   "Carrier_35_PB3_ProdHoldRH" AT %I2117.2 : Bool;   // PB 3 PRODUCTION HOLD RH
   "Carrier_35_PB4_ResetRH" AT %I2117.3 : Bool;   // PB 4 RESET RH
   "Carrier_35_SpareInput(4_14)" AT %I2117.4 : Bool;   // SPARE INPUT
   "Carrier_35_SpareInput(4_15)" AT %I2117.5 : Bool;   // SPARE INPUT
   "Carrier_35_SpareInput(4_16)" AT %I2117.6 : Bool;   // SPARE INPUT
   "Carrier_35_SpareInput(4_17)" AT %I2117.7 : Bool;   // SPARE INPUT
   "Carrier_35_Slot5_Output" AT %IW2118 : Word;   // SLOT 5 OUTPUT WORD
   "Carrier_35_IRD400_HMI_24VDC_ENABLE" AT %I2118.0 : Bool;   // IRD 400 PANEL HMI 24V DC POWER
   "Carrier_35_FaultLight_LH" AT %I2118.1 : Bool;   // FAULT LIGHT LH
   "Carrier_35_RunLight_LH" AT %I2118.2 : Bool;   // RUN LIGHT LH
   "Carrier_35_FaultLight_RH" AT %I2118.3 : Bool;   // FAULT LIGHT RH
   "Carrier_35_RunLight_RH" AT %I2118.4 : Bool;   // RUN LIGHT RH
   "Carrier_35_SpareOutput(5_5)" AT %I2118.5 : Bool;   // SPARE OUTPUT
   "Carrier_35_SpareOutput(5_6)" AT %I2118.6 : Bool;   // SPARE OUTPUT
   "Carrier_35_SpareOutput(5_7)" AT %I2118.7 : Bool;   // SPARE OUTPUT
   "Carrier_35_ActualSpeed" AT %IW2120 : Word;   // ACTUAL SPEED
   "Carrier_35_CarrierDriveAlarm" AT %IW2122 : Word;   // CARRIER DRIVE ALARM
   "Carrier_35_CarrierDriveWarning" AT %IW2124 : Word;   // CARRIER DRIVE WARNING
   "Carrier_36_Status" AT %IW2150 : Word;   // CARRIER STATUS WORD
   "Carrier_36_Status.0" AT %I2150.0 : Bool;   // HEARTBEAT
   "Carrier_36_Status.1" AT %I2150.1 : Bool;   // MANUAL
   "Carrier_36_Status.2" AT %I2150.2 : Bool;   // IN_AUTO
   "Carrier_36_Status.3" AT %I2150.3 : Bool;   // POSITIONING_COMPLETE
   "Carrier_36_Status.4" AT %I2150.4 : Bool;   // PRODUCTION HOLD
   "Carrier_36_Status.5" AT %I2150.5 : Bool;   // CARRIER MOVING FORWARD
   "Carrier_36_Status.6" AT %I2150.6 : Bool;   // CARRIER MOVING REVERSE
   "Carrier_36_Status.7" AT %I2150.7 : Bool;   // CARRIER FAULT
   "Carrier_36_Status.8" AT %I2151.0 : Bool;   // CRASH DETECT TRIPPED
   "Carrier_36_Status.9" AT %I2151.1 : Bool;
   "Carrier_36_Status.10" AT %I2151.2 : Bool;
   "Carrier_36_Status.11" AT %I2151.3 : Bool;
   "Carrier_36_Status.12" AT %I2151.4 : Bool;
   "Carrier_36_Status.13" AT %I2151.5 : Bool;
   "Carrier_36_Status.14" AT %I2151.6 : Bool;
   "Carrier_36_Status.15" AT %I2151.7 : Bool;
   "Carrier_36_SDCFaultCode" AT %IW2152 : Word;   // SDC FAULT CODE
   "Carrier_36_CarrierPosition" AT %ID2154 : DWord;   // CARRIER POSITION
   "Carrier_36_CarrierNumber" AT %IW2158 : Word;   // CARRIER NUMBER
   "Carrier_36_G120DControlWord" AT %IW2160 : Word;   // G120D_STW1_CONTROL
   "Carrier_36_G120DControlWord.0" AT %I2160.0 : Bool;   // Bit_00_ON
   "Carrier_36_G120DControlWord.1" AT %I2160.1 : Bool;   // Bit_01_AUS2_INH
   "Carrier_36_G120DControlWord.2" AT %I2160.2 : Bool;   // Bit_02_AUS3_STOP
   "Carrier_36_G120DControlWord.3" AT %I2160.3 : Bool;   // Bit_03_EN
   "Carrier_36_G120DControlWord.4" AT %I2160.4 : Bool;   // Bit_04_EN_RAMP
   "Carrier_36_G120DControlWord.5" AT %I2160.5 : Bool;   // Bit_05_START_RAMP
   "Carrier_36_G120DControlWord.6" AT %I2160.6 : Bool;   // Bit_06_SETPOINT
   "Carrier_36_G120DControlWord.7" AT %I2160.7 : Bool;   // Bit_07_RESET
   "Carrier_36_G120DControlWord.8" AT %I2161.0 : Bool;   // Bit_08_JOG_R
   "Carrier_36_G120DControlWord.9" AT %I2161.1 : Bool;   // Bit_09_JOG_L
   "Carrier_36_G120DControlWord.10" AT %I2161.2 : Bool;   // Bit_10_CONTR_PLC
   "Carrier_36_G120DControlWord.11" AT %I2161.3 : Bool;   // Bit_11_REVERSE
   "Carrier_36_G120DControlWord.12" AT %I2161.4 : Bool;   // Bit_12_BRAKE_RELEASE
   "Carrier_36_G120DControlWord.13" AT %I2161.5 : Bool;   // Bit_13_DDS
   "Carrier_36_G120DControlWord.14" AT %I2161.6 : Bool;   // Bit_14_DO0
   "Carrier_36_G120DControlWord.15" AT %I2161.7 : Bool;   // Bit_15_DO1
   "Carrier_36_G120DStatusWord" AT %IW2162 : Word;   // G120D_ZSW1_STATUS
   "Carrier_36_G120DStatusWord.0" AT %I2162.0 : Bool;   // Bit_00_READY_RUN
   "Carrier_36_G120DStatusWord.1" AT %I2162.1 : Bool;   // Bit_01_READY_ON
   "Carrier_36_G120DStatusWord.2" AT %I2162.2 : Bool;   // Bit_02_ENABLE
   "Carrier_36_G120DStatusWord.3" AT %I2162.3 : Bool;   // Bit_03_FAULT
   "Carrier_36_G120DStatusWord.4" AT %I2162.4 : Bool;   // Bit_04_OFF2
   "Carrier_36_G120DStatusWord.5" AT %I2162.5 : Bool;   // Bit_05_OFF3
   "Carrier_36_G120DStatusWord.6" AT %I2162.6 : Bool;   // Bit_06_LOCK_OUT
   "Carrier_36_G120DStatusWord.7" AT %I2162.7 : Bool;   // Bit_07_WARN
   "Carrier_36_G120DStatusWord.8" AT %I2163.0 : Bool;   // Bit_08_NO_DEVIATION
   "Carrier_36_G120DStatusWord.9" AT %I2163.1 : Bool;   // Bit_09_CONTR_PLC
   "Carrier_36_G120DStatusWord.10" AT %I2163.2 : Bool;   // Bit_10_F_MAX
   "Carrier_36_G120DStatusWord.11" AT %I2163.3 : Bool;   // Bit_11_LIMIT_REACHED
   "Carrier_36_G120DStatusWord.12" AT %I2163.4 : Bool;   // Bit_12_BRAKE_OPEN
   "Carrier_36_G120DStatusWord.13" AT %I2163.5 : Bool;   // Bit_13_NO_OVERTEMP
   "Carrier_36_G120DStatusWord.14" AT %I2163.6 : Bool;   // Bit_14_CW_CCW
   "Carrier_36_G120DStatusWord.15" AT %I2163.7 : Bool;   // Bit_15_OVERL
   "Carrier_36_Slot2_Input" AT %IW2164 : Word;   // SLOT 2 INPUT WORD
   "Carrier_36_CrashDetectSW" AT %I2164.0 : Bool;   // CRASH DETECT SW
   "Carrier_36_SpareSafetyInput(2_1)" AT %I2164.1 : Bool;   // SPARE SAFETY INPUT
   "Carrier_36_SpareSafetyInput(2_2)" AT %I2164.2 : Bool;   // SPARE SAFETY INPUT
   "Carrier_36_SpareSafetyInput(2_3)" AT %I2164.3 : Bool;   // SPARE SAFETY INPUT
   "Carrier_36_SpareSafetyInput(2_4)" AT %I2164.4 : Bool;   // SPARE SAFETY INPUT
   "Carrier_36_SpareSafetyInput(2_5)" AT %I2164.5 : Bool;   // SPARE SAFETY INPUT
   "Carrier_36_SpareSafetyInput(2_6)" AT %I2164.6 : Bool;   // SPARE SAFETY INPUT
   "Carrier_36_SpareSafetyInput(2_7)" AT %I2164.7 : Bool;   // SPARE SAFETY INPUT
   "Carrier_36_Slot3_SafetyOutput" AT %IW2165 : Word;   // SLOT 3 SAFETY OUTPUT WORD
   "Carrier_36_Crash_Detect_OK" AT %I2165.0 : Bool;   // CARRIER CRASH DETECT
   "Carrier_36_SpareSafetyOutput(3_1)" AT %I2165.1 : Bool;   // SPARE SAFETY OUTPUT
   "Carrier_36_SpareSafetyOutput(3_2)" AT %I2165.2 : Bool;   // SPARE SAFETY OUTPUT
   "Carrier_36_SpareSafetyOutput(3_3)" AT %I2165.3 : Bool;   // SPARE SAFETY OUTPUT
   "Carrier_36_SpareSafetyOutput(3_4)" AT %I2165.4 : Bool;   // SPARE SAFETY OUTPUT
   "Carrier_36_SpareSafetyOutput(3_5)" AT %I2165.5 : Bool;   // SPARE SAFETY OUTPUT
   "Carrier_36_SpareSafetyOutput(3_6)" AT %I2165.6 : Bool;   // SPARE SAFETY OUTPUT
   "Carrier_36_SpareSafetyOutput(3_7)" AT %I2165.7 : Bool;   // SPARE SAFETY OUTPUT
   "Carrier_36_Slot4_Input" AT %IW2166 : Word;   // SLOT 4 INPUT WORD
   "Carrier_36_480VPowerOn_MDCB1" AT %I2166.0 : Bool;   // 480 VAC POWER ON MDCB 1
   "Carrier_36_SpareInput(4_1)" AT %I2166.1 : Bool;   // SPARE INPUT
   "Carrier_36_SpareInput(4_2)" AT %I2166.2 : Bool;   // SPARE INPUT
   "Carrier_36_SitopSelectStatus" AT %I2166.3 : Bool;   // SITOP SELECT STATUS
   "Carrier_36_DCsupplyOnPSCB2" AT %I2166.4 : Bool;   // DC SUPPLY ON PSCB 2
   "Carrier_36_SpareInput(4_5)" AT %I2166.5 : Bool;   // SPARE INPUT
   "Carrier_36_SpareInput(4_6)" AT %I2166.6 : Bool;   // SPARE INPUT
   "Carrier_36_SpareInput(4_7)" AT %I2166.7 : Bool;   // SPARE INPUT
   "Carrier_36_PB1_ProdHoldLH" AT %I2167.0 : Bool;   // PB 1 PRODUCTION HOLD LH
   "Carrier_36_PB2_ResetLH" AT %I2167.1 : Bool;   // PB 2 RESET LH
   "Carrier_36_PB3_ProdHoldRH" AT %I2167.2 : Bool;   // PB 3 PRODUCTION HOLD RH
   "Carrier_36_PB4_ResetRH" AT %I2167.3 : Bool;   // PB 4 RESET RH
   "Carrier_36_SpareInput(4_14)" AT %I2167.4 : Bool;   // SPARE INPUT
   "Carrier_36_SpareInput(4_15)" AT %I2167.5 : Bool;   // SPARE INPUT
   "Carrier_36_SpareInput(4_16)" AT %I2167.6 : Bool;   // SPARE INPUT
   "Carrier_36_SpareInput(4_17)" AT %I2167.7 : Bool;   // SPARE INPUT
   "Carrier_36_Slot5_Output" AT %IW2168 : Word;   // SLOT 5 OUTPUT WORD
   "Carrier_36_IRD400_HMI_24VDC_ENABLE" AT %I2168.0 : Bool;   // IRD 400 PANEL HMI 24V DC POWER
   "Carrier_36_FaultLight_LH" AT %I2168.1 : Bool;   // FAULT LIGHT LH
   "Carrier_36_RunLight_LH" AT %I2168.2 : Bool;   // RUN LIGHT LH
   "Carrier_36_FaultLight_RH" AT %I2168.3 : Bool;   // FAULT LIGHT RH
   "Carrier_36_RunLight_RH" AT %I2168.4 : Bool;   // RUN LIGHT RH
   "Carrier_36_SpareOutput(5_5)" AT %I2168.5 : Bool;   // SPARE OUTPUT
   "Carrier_36_SpareOutput(5_6)" AT %I2168.6 : Bool;   // SPARE OUTPUT
   "Carrier_36_SpareOutput(5_7)" AT %I2168.7 : Bool;   // SPARE OUTPUT
   "Carrier_36_ActualSpeed" AT %IW2170 : Word;   // ACTUAL SPEED
   "Carrier_36_CarrierDriveAlarm" AT %IW2172 : Word;   // CARRIER DRIVE ALARM
   "Carrier_36_CarrierDriveWarning" AT %IW2174 : Word;   // CARRIER DRIVE WARNING
   "Carrier_37_Status" AT %IW2200 : Word;   // CARRIER STATUS WORD
   "Carrier_37_Status.0" AT %I2200.0 : Bool;   // HEARTBEAT
   "Carrier_37_Status.1" AT %I2200.1 : Bool;   // MANUAL
   "Carrier_37_Status.2" AT %I2200.2 : Bool;   // IN_AUTO
   "Carrier_37_Status.3" AT %I2200.3 : Bool;   // POSITIONING_COMPLETE
   "Carrier_37_Status.4" AT %I2200.4 : Bool;   // PRODUCTION HOLD
   "Carrier_37_Status.5" AT %I2200.5 : Bool;   // CARRIER MOVING FORWARD
   "Carrier_37_Status.6" AT %I2200.6 : Bool;   // CARRIER MOVING REVERSE
   "Carrier_37_Status.7" AT %I2200.7 : Bool;   // CARRIER FAULT
   "Carrier_37_Status.8" AT %I2201.0 : Bool;   // CRASH DETECT TRIPPED
   "Carrier_37_Status.9" AT %I2201.1 : Bool;
   "Carrier_37_Status.10" AT %I2201.2 : Bool;
   "Carrier_37_Status.11" AT %I2201.3 : Bool;
   "Carrier_37_Status.12" AT %I2201.4 : Bool;
   "Carrier_37_Status.13" AT %I2201.5 : Bool;
   "Carrier_37_Status.14" AT %I2201.6 : Bool;
   "Carrier_37_Status.15" AT %I2201.7 : Bool;
   "Carrier_37_SDCFaultCode" AT %IW2202 : Word;   // SDC FAULT CODE
   "Carrier_37_CarrierPosition" AT %ID2204 : DWord;   // CARRIER POSITION
   "Carrier_37_CarrierNumber" AT %IW2208 : Word;   // CARRIER NUMBER
   "Carrier_37_G120DControlWord" AT %IW2210 : Word;   // G120D_STW1_CONTROL
   "Carrier_37_G120DControlWord.0" AT %I2210.0 : Bool;   // Bit_00_ON
   "Carrier_37_G120DControlWord.1" AT %I2210.1 : Bool;   // Bit_01_AUS2_INH
   "Carrier_37_G120DControlWord.2" AT %I2210.2 : Bool;   // Bit_02_AUS3_STOP
   "Carrier_37_G120DControlWord.3" AT %I2210.3 : Bool;   // Bit_03_EN
   "Carrier_37_G120DControlWord.4" AT %I2210.4 : Bool;   // Bit_04_EN_RAMP
   "Carrier_37_G120DControlWord.5" AT %I2210.5 : Bool;   // Bit_05_START_RAMP
   "Carrier_37_G120DControlWord.6" AT %I2210.6 : Bool;   // Bit_06_SETPOINT
   "Carrier_37_G120DControlWord.7" AT %I2210.7 : Bool;   // Bit_07_RESET
   "Carrier_37_G120DControlWord.8" AT %I2211.0 : Bool;   // Bit_08_JOG_R
   "Carrier_37_G120DControlWord.9" AT %I2211.1 : Bool;   // Bit_09_JOG_L
   "Carrier_37_G120DControlWord.10" AT %I2211.2 : Bool;   // Bit_10_CONTR_PLC
   "Carrier_37_G120DControlWord.11" AT %I2211.3 : Bool;   // Bit_11_REVERSE
   "Carrier_37_G120DControlWord.12" AT %I2211.4 : Bool;   // Bit_12_BRAKE_RELEASE
   "Carrier_37_G120DControlWord.13" AT %I2211.5 : Bool;   // Bit_13_DDS
   "Carrier_37_G120DControlWord.14" AT %I2211.6 : Bool;   // Bit_14_DO0
   "Carrier_37_G120DControlWord.15" AT %I2211.7 : Bool;   // Bit_15_DO1
   "Carrier_37_G120DStatusWord" AT %IW2212 : Word;   // G120D_ZSW1_STATUS
   "Carrier_37_G120DStatusWord.0" AT %I2212.0 : Bool;   // Bit_00_READY_RUN
   "Carrier_37_G120DStatusWord.1" AT %I2212.1 : Bool;   // Bit_01_READY_ON
   "Carrier_37_G120DStatusWord.2" AT %I2212.2 : Bool;   // Bit_02_ENABLE
   "Carrier_37_G120DStatusWord.3" AT %I2212.3 : Bool;   // Bit_03_FAULT
   "Carrier_37_G120DStatusWord.4" AT %I2212.4 : Bool;   // Bit_04_OFF2
   "Carrier_37_G120DStatusWord.5" AT %I2212.5 : Bool;   // Bit_05_OFF3
   "Carrier_37_G120DStatusWord.6" AT %I2212.6 : Bool;   // Bit_06_LOCK_OUT
   "Carrier_37_G120DStatusWord.7" AT %I2212.7 : Bool;   // Bit_07_WARN
   "Carrier_37_G120DStatusWord.8" AT %I2213.0 : Bool;   // Bit_08_NO_DEVIATION
   "Carrier_37_G120DStatusWord.9" AT %I2213.1 : Bool;   // Bit_09_CONTR_PLC
   "Carrier_37_G120DStatusWord.10" AT %I2213.2 : Bool;   // Bit_10_F_MAX
   "Carrier_37_G120DStatusWord.11" AT %I2213.3 : Bool;   // Bit_11_LIMIT_REACHED
   "Carrier_37_G120DStatusWord.12" AT %I2213.4 : Bool;   // Bit_12_BRAKE_OPEN
   "Carrier_37_G120DStatusWord.13" AT %I2213.5 : Bool;   // Bit_13_NO_OVERTEMP
   "Carrier_37_G120DStatusWord.14" AT %I2213.6 : Bool;   // Bit_14_CW_CCW
   "Carrier_37_G120DStatusWord.15" AT %I2213.7 : Bool;   // Bit_15_OVERL
   "Carrier_37_Slot2_Input" AT %IW2214 : Word;   // SLOT 2 INPUT WORD
   "Carrier_37_CrashDetectSW" AT %I2214.0 : Bool;   // CRASH DETECT SW
   "Carrier_37_SpareSafetyInput(2_1)" AT %I2214.1 : Bool;   // SPARE SAFETY INPUT
   "Carrier_37_SpareSafetyInput(2_2)" AT %I2214.2 : Bool;   // SPARE SAFETY INPUT
   "Carrier_37_SpareSafetyInput(2_3)" AT %I2214.3 : Bool;   // SPARE SAFETY INPUT
   "Carrier_37_SpareSafetyInput(2_4)" AT %I2214.4 : Bool;   // SPARE SAFETY INPUT
   "Carrier_37_SpareSafetyInput(2_5)" AT %I2214.5 : Bool;   // SPARE SAFETY INPUT
   "Carrier_37_SpareSafetyInput(2_6)" AT %I2214.6 : Bool;   // SPARE SAFETY INPUT
   "Carrier_37_SpareSafetyInput(2_7)" AT %I2214.7 : Bool;   // SPARE SAFETY INPUT
   "Carrier_37_Slot3_SafetyOutput" AT %IW2215 : Word;   // SLOT 3 SAFETY OUTPUT WORD
   "Carrier_37_Crash_Detect_OK" AT %I2215.0 : Bool;   // CARRIER CRASH DETECT
   "Carrier_37_SpareSafetyOutput(3_1)" AT %I2215.1 : Bool;   // SPARE SAFETY OUTPUT
   "Carrier_37_SpareSafetyOutput(3_2)" AT %I2215.2 : Bool;   // SPARE SAFETY OUTPUT
   "Carrier_37_SpareSafetyOutput(3_3)" AT %I2215.3 : Bool;   // SPARE SAFETY OUTPUT
   "Carrier_37_SpareSafetyOutput(3_4)" AT %I2215.4 : Bool;   // SPARE SAFETY OUTPUT
   "Carrier_37_SpareSafetyOutput(3_5)" AT %I2215.5 : Bool;   // SPARE SAFETY OUTPUT
   "Carrier_37_SpareSafetyOutput(3_6)" AT %I2215.6 : Bool;   // SPARE SAFETY OUTPUT
   "Carrier_37_SpareSafetyOutput(3_7)" AT %I2215.7 : Bool;   // SPARE SAFETY OUTPUT
   "Carrier_37_Slot4_Input" AT %IW2216 : Word;   // SLOT 4 INPUT WORD
   "Carrier_37_480VPowerOn_MDCB1" AT %I2216.0 : Bool;   // 480 VAC POWER ON MDCB 1
   "Carrier_37_SpareInput(4_1)" AT %I2216.1 : Bool;   // SPARE INPUT
   "Carrier_37_SpareInput(4_2)" AT %I2216.2 : Bool;   // SPARE INPUT
   "Carrier_37_SitopSelectStatus" AT %I2216.3 : Bool;   // SITOP SELECT STATUS
   "Carrier_37_DCsupplyOnPSCB2" AT %I2216.4 : Bool;   // DC SUPPLY ON PSCB 2
   "Carrier_37_SpareInput(4_5)" AT %I2216.5 : Bool;   // SPARE INPUT
   "Carrier_37_SpareInput(4_6)" AT %I2216.6 : Bool;   // SPARE INPUT
   "Carrier_37_SpareInput(4_7)" AT %I2216.7 : Bool;   // SPARE INPUT
   "Carrier_37_PB1_ProdHoldLH" AT %I2217.0 : Bool;   // PB 1 PRODUCTION HOLD LH
   "Carrier_37_PB2_ResetLH" AT %I2217.1 : Bool;   // PB 2 RESET LH
   "Carrier_37_PB3_ProdHoldRH" AT %I2217.2 : Bool;   // PB 3 PRODUCTION HOLD RH
   "Carrier_37_PB4_ResetRH" AT %I2217.3 : Bool;   // PB 4 RESET RH
   "Carrier_37_SpareInput(4_14)" AT %I2217.4 : Bool;   // SPARE INPUT
   "Carrier_37_SpareInput(4_15)" AT %I2217.5 : Bool;   // SPARE INPUT
   "Carrier_37_SpareInput(4_16)" AT %I2217.6 : Bool;   // SPARE INPUT
   "Carrier_37_SpareInput(4_17)" AT %I2217.7 : Bool;   // SPARE INPUT
   "Carrier_37_Slot5_Output" AT %IW2218 : Word;   // SLOT 5 OUTPUT WORD
   "Carrier_37_IRD400_HMI_24VDC_ENABLE" AT %I2218.0 : Bool;   // IRD 400 PANEL HMI 24V DC POWER
   "Carrier_37_FaultLight_LH" AT %I2218.1 : Bool;   // FAULT LIGHT LH
   "Carrier_37_RunLight_LH" AT %I2218.2 : Bool;   // RUN LIGHT LH
   "Carrier_37_FaultLight_RH" AT %I2218.3 : Bool;   // FAULT LIGHT RH
   "Carrier_37_RunLight_RH" AT %I2218.4 : Bool;   // RUN LIGHT RH
   "Carrier_37_SpareOutput(5_5)" AT %I2218.5 : Bool;   // SPARE OUTPUT
   "Carrier_37_SpareOutput(5_6)" AT %I2218.6 : Bool;   // SPARE OUTPUT
   "Carrier_37_SpareOutput(5_7)" AT %I2218.7 : Bool;   // SPARE OUTPUT
   "Carrier_37_ActualSpeed" AT %IW2220 : Word;   // ACTUAL SPEED
   "Carrier_37_CarrierDriveAlarm" AT %IW2222 : Word;   // CARRIER DRIVE ALARM
   "Carrier_37_CarrierDriveWarning" AT %IW2224 : Word;   // CARRIER DRIVE WARNING
   "Carrier_38_Status" AT %IW2250 : Word;   // CARRIER STATUS WORD
   "Carrier_38_Status.0" AT %I2250.0 : Bool;   // HEARTBEAT
   "Carrier_38_Status.1" AT %I2250.1 : Bool;   // MANUAL
   "Carrier_38_Status.2" AT %I2250.2 : Bool;   // IN_AUTO
   "Carrier_38_Status.3" AT %I2250.3 : Bool;   // POSITIONING_COMPLETE
   "Carrier_38_Status.4" AT %I2250.4 : Bool;   // PRODUCTION HOLD
   "Carrier_38_Status.5" AT %I2250.5 : Bool;   // CARRIER MOVING FORWARD
   "Carrier_38_Status.6" AT %I2250.6 : Bool;   // CARRIER MOVING REVERSE
   "Carrier_38_Status.7" AT %I2250.7 : Bool;   // CARRIER FAULT
   "Carrier_38_Status.8" AT %I2251.0 : Bool;   // CRASH DETECT TRIPPED
   "Carrier_38_Status.9" AT %I2251.1 : Bool;
   "Carrier_38_Status.10" AT %I2251.2 : Bool;
   "Carrier_38_Status.11" AT %I2251.3 : Bool;
   "Carrier_38_Status.12" AT %I2251.4 : Bool;
   "Carrier_38_Status.13" AT %I2251.5 : Bool;
   "Carrier_38_Status.14" AT %I2251.6 : Bool;
   "Carrier_38_Status.15" AT %I2251.7 : Bool;
   "Carrier_38_SDCFaultCode" AT %IW2252 : Word;   // SDC FAULT CODE
   "Carrier_38_CarrierPosition" AT %ID2254 : DWord;   // CARRIER POSITION
   "Carrier_38_CarrierNumber" AT %IW2258 : Word;   // CARRIER NUMBER
   "Carrier_38_G120DControlWord" AT %IW2260 : Word;   // G120D_STW1_CONTROL
   "Carrier_38_G120DControlWord.0" AT %I2260.0 : Bool;   // Bit_00_ON
   "Carrier_38_G120DControlWord.1" AT %I2260.1 : Bool;   // Bit_01_AUS2_INH
   "Carrier_38_G120DControlWord.2" AT %I2260.2 : Bool;   // Bit_02_AUS3_STOP
   "Carrier_38_G120DControlWord.3" AT %I2260.3 : Bool;   // Bit_03_EN
   "Carrier_38_G120DControlWord.4" AT %I2260.4 : Bool;   // Bit_04_EN_RAMP
   "Carrier_38_G120DControlWord.5" AT %I2260.5 : Bool;   // Bit_05_START_RAMP
   "Carrier_38_G120DControlWord.6" AT %I2260.6 : Bool;   // Bit_06_SETPOINT
   "Carrier_38_G120DControlWord.7" AT %I2260.7 : Bool;   // Bit_07_RESET
   "Carrier_38_G120DControlWord.8" AT %I2261.0 : Bool;   // Bit_08_JOG_R
   "Carrier_38_G120DControlWord.9" AT %I2261.1 : Bool;   // Bit_09_JOG_L
   "Carrier_38_G120DControlWord.10" AT %I2261.2 : Bool;   // Bit_10_CONTR_PLC
   "Carrier_38_G120DControlWord.11" AT %I2261.3 : Bool;   // Bit_11_REVERSE
   "Carrier_38_G120DControlWord.12" AT %I2261.4 : Bool;   // Bit_12_BRAKE_RELEASE
   "Carrier_38_G120DControlWord.13" AT %I2261.5 : Bool;   // Bit_13_DDS
   "Carrier_38_G120DControlWord.14" AT %I2261.6 : Bool;   // Bit_14_DO0
   "Carrier_38_G120DControlWord.15" AT %I2261.7 : Bool;   // Bit_15_DO1
   "Carrier_38_G120DStatusWord" AT %IW2262 : Word;   // G120D_ZSW1_STATUS
   "Carrier_38_G120DStatusWord.0" AT %I2262.0 : Bool;   // Bit_00_READY_RUN
   "Carrier_38_G120DStatusWord.1" AT %I2262.1 : Bool;   // Bit_01_READY_ON
   "Carrier_38_G120DStatusWord.2" AT %I2262.2 : Bool;   // Bit_02_ENABLE
   "Carrier_38_G120DStatusWord.3" AT %I2262.3 : Bool;   // Bit_03_FAULT
   "Carrier_38_G120DStatusWord.4" AT %I2262.4 : Bool;   // Bit_04_OFF2
   "Carrier_38_G120DStatusWord.5" AT %I2262.5 : Bool;   // Bit_05_OFF3
   "Carrier_38_G120DStatusWord.6" AT %I2262.6 : Bool;   // Bit_06_LOCK_OUT
   "Carrier_38_G120DStatusWord.7" AT %I2262.7 : Bool;   // Bit_07_WARN
   "Carrier_38_G120DStatusWord.8" AT %I2263.0 : Bool;   // Bit_08_NO_DEVIATION
   "Carrier_38_G120DStatusWord.9" AT %I2263.1 : Bool;   // Bit_09_CONTR_PLC
   "Carrier_38_G120DStatusWord.10" AT %I2263.2 : Bool;   // Bit_10_F_MAX
   "Carrier_38_G120DStatusWord.11" AT %I2263.3 : Bool;   // Bit_11_LIMIT_REACHED
   "Carrier_38_G120DStatusWord.12" AT %I2263.4 : Bool;   // Bit_12_BRAKE_OPEN
   "Carrier_38_G120DStatusWord.13" AT %I2263.5 : Bool;   // Bit_13_NO_OVERTEMP
   "Carrier_38_G120DStatusWord.14" AT %I2263.6 : Bool;   // Bit_14_CW_CCW
   "Carrier_38_G120DStatusWord.15" AT %I2263.7 : Bool;   // Bit_15_OVERL
   "Carrier_38_Slot2_Input" AT %IW2264 : Word;   // SLOT 2 INPUT WORD
   "Carrier_38_CrashDetectSW" AT %I2264.0 : Bool;   // CRASH DETECT SW
   "Carrier_38_SpareSafetyInput(2_1)" AT %I2264.1 : Bool;   // SPARE SAFETY INPUT
   "Carrier_38_SpareSafetyInput(2_2)" AT %I2264.2 : Bool;   // SPARE SAFETY INPUT
   "Carrier_38_SpareSafetyInput(2_3)" AT %I2264.3 : Bool;   // SPARE SAFETY INPUT
   "Carrier_38_SpareSafetyInput(2_4)" AT %I2264.4 : Bool;   // SPARE SAFETY INPUT
   "Carrier_38_SpareSafetyInput(2_5)" AT %I2264.5 : Bool;   // SPARE SAFETY INPUT
   "Carrier_38_SpareSafetyInput(2_6)" AT %I2264.6 : Bool;   // SPARE SAFETY INPUT
   "Carrier_38_SpareSafetyInput(2_7)" AT %I2264.7 : Bool;   // SPARE SAFETY INPUT
   "Carrier_38_Slot3_SafetyOutput" AT %IW2265 : Word;   // SLOT 3 SAFETY OUTPUT WORD
   "Carrier_38_Crash_Detect_OK" AT %I2265.0 : Bool;   // CARRIER CRASH DETECT
   "Carrier_38_SpareSafetyOutput(3_1)" AT %I2265.1 : Bool;   // SPARE SAFETY OUTPUT
   "Carrier_38_SpareSafetyOutput(3_2)" AT %I2265.2 : Bool;   // SPARE SAFETY OUTPUT
   "Carrier_38_SpareSafetyOutput(3_3)" AT %I2265.3 : Bool;   // SPARE SAFETY OUTPUT
   "Carrier_38_SpareSafetyOutput(3_4)" AT %I2265.4 : Bool;   // SPARE SAFETY OUTPUT
   "Carrier_38_SpareSafetyOutput(3_5)" AT %I2265.5 : Bool;   // SPARE SAFETY OUTPUT
   "Carrier_38_SpareSafetyOutput(3_6)" AT %I2265.6 : Bool;   // SPARE SAFETY OUTPUT
   "Carrier_38_SpareSafetyOutput(3_7)" AT %I2265.7 : Bool;   // SPARE SAFETY OUTPUT
   "Carrier_38_Slot4_Input" AT %IW2266 : Word;   // SLOT 4 INPUT WORD
   "Carrier_38_480VPowerOn_MDCB1" AT %I2266.0 : Bool;   // 480 VAC POWER ON MDCB 1
   "Carrier_38_SpareInput(4_1)" AT %I2266.1 : Bool;   // SPARE INPUT
   "Carrier_38_SpareInput(4_2)" AT %I2266.2 : Bool;   // SPARE INPUT
   "Carrier_38_SitopSelectStatus" AT %I2266.3 : Bool;   // SITOP SELECT STATUS
   "Carrier_38_DCsupplyOnPSCB2" AT %I2266.4 : Bool;   // DC SUPPLY ON PSCB 2
   "Carrier_38_SpareInput(4_5)" AT %I2266.5 : Bool;   // SPARE INPUT
   "Carrier_38_SpareInput(4_6)" AT %I2266.6 : Bool;   // SPARE INPUT
   "Carrier_38_SpareInput(4_7)" AT %I2266.7 : Bool;   // SPARE INPUT
   "Carrier_38_PB1_ProdHoldLH" AT %I2267.0 : Bool;   // PB 1 PRODUCTION HOLD LH
   "Carrier_38_PB2_ResetLH" AT %I2267.1 : Bool;   // PB 2 RESET LH
   "Carrier_38_PB3_ProdHoldRH" AT %I2267.2 : Bool;   // PB 3 PRODUCTION HOLD RH
   "Carrier_38_PB4_ResetRH" AT %I2267.3 : Bool;   // PB 4 RESET RH
   "Carrier_38_SpareInput(4_14)" AT %I2267.4 : Bool;   // SPARE INPUT
   "Carrier_38_SpareInput(4_15)" AT %I2267.5 : Bool;   // SPARE INPUT
   "Carrier_38_SpareInput(4_16)" AT %I2267.6 : Bool;   // SPARE INPUT
   "Carrier_38_SpareInput(4_17)" AT %I2267.7 : Bool;   // SPARE INPUT
   "Carrier_38_Slot5_Output" AT %IW2268 : Word;   // SLOT 5 OUTPUT WORD
   "Carrier_38_IRD400_HMI_24VDC_ENABLE" AT %I2268.0 : Bool;   // IRD 400 PANEL HMI 24V DC POWER
   "Carrier_38_FaultLight_LH" AT %I2268.1 : Bool;   // FAULT LIGHT LH
   "Carrier_38_RunLight_LH" AT %I2268.2 : Bool;   // RUN LIGHT LH
   "Carrier_38_FaultLight_RH" AT %I2268.3 : Bool;   // FAULT LIGHT RH
   "Carrier_38_RunLight_RH" AT %I2268.4 : Bool;   // RUN LIGHT RH
   "Carrier_38_SpareOutput(5_5)" AT %I2268.5 : Bool;   // SPARE OUTPUT
   "Carrier_38_SpareOutput(5_6)" AT %I2268.6 : Bool;   // SPARE OUTPUT
   "Carrier_38_SpareOutput(5_7)" AT %I2268.7 : Bool;   // SPARE OUTPUT
   "Carrier_38_ActualSpeed" AT %IW2270 : Word;   // ACTUAL SPEED
   "Carrier_38_CarrierDriveAlarm" AT %IW2272 : Word;   // CARRIER DRIVE ALARM
   "Carrier_38_CarrierDriveWarning" AT %IW2274 : Word;   // CARRIER DRIVE WARNING
   "Carrier_39_Status" AT %IW2300 : Word;   // CARRIER STATUS WORD
   "Carrier_39_Status.0" AT %I2300.0 : Bool;   // HEARTBEAT
   "Carrier_39_Status.1" AT %I2300.1 : Bool;   // MANUAL
   "Carrier_39_Status.2" AT %I2300.2 : Bool;   // IN_AUTO
   "Carrier_39_Status.3" AT %I2300.3 : Bool;   // POSITIONING_COMPLETE
   "Carrier_39_Status.4" AT %I2300.4 : Bool;   // PRODUCTION HOLD
   "Carrier_39_Status.5" AT %I2300.5 : Bool;   // CARRIER MOVING FORWARD
   "Carrier_39_Status.6" AT %I2300.6 : Bool;   // CARRIER MOVING REVERSE
   "Carrier_39_Status.7" AT %I2300.7 : Bool;   // CARRIER FAULT
   "Carrier_39_Status.8" AT %I2301.0 : Bool;   // CRASH DETECT TRIPPED
   "Carrier_39_Status.9" AT %I2301.1 : Bool;
   "Carrier_39_Status.10" AT %I2301.2 : Bool;
   "Carrier_39_Status.11" AT %I2301.3 : Bool;
   "Carrier_39_Status.12" AT %I2301.4 : Bool;
   "Carrier_39_Status.13" AT %I2301.5 : Bool;
   "Carrier_39_Status.14" AT %I2301.6 : Bool;
   "Carrier_39_Status.15" AT %I2301.7 : Bool;
   "Carrier_39_SDCFaultCode" AT %IW2302 : Word;   // SDC FAULT CODE
   "Carrier_39_CarrierPosition" AT %ID2304 : DWord;   // CARRIER POSITION
   "Carrier_39_CarrierNumber" AT %IW2308 : Word;   // CARRIER NUMBER
   "Carrier_39_G120DControlWord" AT %IW2310 : Word;   // G120D_STW1_CONTROL
   "Carrier_39_G120DControlWord.0" AT %I2310.0 : Bool;   // Bit_00_ON
   "Carrier_39_G120DControlWord.1" AT %I2310.1 : Bool;   // Bit_01_AUS2_INH
   "Carrier_39_G120DControlWord.2" AT %I2310.2 : Bool;   // Bit_02_AUS3_STOP
   "Carrier_39_G120DControlWord.3" AT %I2310.3 : Bool;   // Bit_03_EN
   "Carrier_39_G120DControlWord.4" AT %I2310.4 : Bool;   // Bit_04_EN_RAMP
   "Carrier_39_G120DControlWord.5" AT %I2310.5 : Bool;   // Bit_05_START_RAMP
   "Carrier_39_G120DControlWord.6" AT %I2310.6 : Bool;   // Bit_06_SETPOINT
   "Carrier_39_G120DControlWord.7" AT %I2310.7 : Bool;   // Bit_07_RESET
   "Carrier_39_G120DControlWord.8" AT %I2311.0 : Bool;   // Bit_08_JOG_R
   "Carrier_39_G120DControlWord.9" AT %I2311.1 : Bool;   // Bit_09_JOG_L
   "Carrier_39_G120DControlWord.10" AT %I2311.2 : Bool;   // Bit_10_CONTR_PLC
   "Carrier_39_G120DControlWord.11" AT %I2311.3 : Bool;   // Bit_11_REVERSE
   "Carrier_39_G120DControlWord.12" AT %I2311.4 : Bool;   // Bit_12_BRAKE_RELEASE
   "Carrier_39_G120DControlWord.13" AT %I2311.5 : Bool;   // Bit_13_DDS
   "Carrier_39_G120DControlWord.14" AT %I2311.6 : Bool;   // Bit_14_DO0
   "Carrier_39_G120DControlWord.15" AT %I2311.7 : Bool;   // Bit_15_DO1
   "Carrier_39_G120DStatusWord" AT %IW2312 : Word;   // G120D_ZSW1_STATUS
   "Carrier_39_G120DStatusWord.0" AT %I2312.0 : Bool;   // Bit_00_READY_RUN
   "Carrier_39_G120DStatusWord.1" AT %I2312.1 : Bool;   // Bit_01_READY_ON
   "Carrier_39_G120DStatusWord.2" AT %I2312.2 : Bool;   // Bit_02_ENABLE
   "Carrier_39_G120DStatusWord.3" AT %I2312.3 : Bool;   // Bit_03_FAULT
   "Carrier_39_G120DStatusWord.4" AT %I2312.4 : Bool;   // Bit_04_OFF2
   "Carrier_39_G120DStatusWord.5" AT %I2312.5 : Bool;   // Bit_05_OFF3
   "Carrier_39_G120DStatusWord.6" AT %I2312.6 : Bool;   // Bit_06_LOCK_OUT
   "Carrier_39_G120DStatusWord.7" AT %I2312.7 : Bool;   // Bit_07_WARN
   "Carrier_39_G120DStatusWord.8" AT %I2313.0 : Bool;   // Bit_08_NO_DEVIATION
   "Carrier_39_G120DStatusWord.9" AT %I2313.1 : Bool;   // Bit_09_CONTR_PLC
   "Carrier_39_G120DStatusWord.10" AT %I2313.2 : Bool;   // Bit_10_F_MAX
   "Carrier_39_G120DStatusWord.11" AT %I2313.3 : Bool;   // Bit_11_LIMIT_REACHED
   "Carrier_39_G120DStatusWord.12" AT %I2313.4 : Bool;   // Bit_12_BRAKE_OPEN
   "Carrier_39_G120DStatusWord.13" AT %I2313.5 : Bool;   // Bit_13_NO_OVERTEMP
   "Carrier_39_G120DStatusWord.14" AT %I2313.6 : Bool;   // Bit_14_CW_CCW
   "Carrier_39_G120DStatusWord.15" AT %I2313.7 : Bool;   // Bit_15_OVERL
   "Carrier_39_Slot2_Input" AT %IW2314 : Word;   // SLOT 2 INPUT WORD
   "Carrier_39_CrashDetectSW" AT %I2314.0 : Bool;   // CRASH DETECT SW
   "Carrier_39_SpareSafetyInput(2_1)" AT %I2314.1 : Bool;   // SPARE SAFETY INPUT
   "Carrier_39_SpareSafetyInput(2_2)" AT %I2314.2 : Bool;   // SPARE SAFETY INPUT
   "Carrier_39_SpareSafetyInput(2_3)" AT %I2314.3 : Bool;   // SPARE SAFETY INPUT
   "Carrier_39_SpareSafetyInput(2_4)" AT %I2314.4 : Bool;   // SPARE SAFETY INPUT
   "Carrier_39_SpareSafetyInput(2_5)" AT %I2314.5 : Bool;   // SPARE SAFETY INPUT
   "Carrier_39_SpareSafetyInput(2_6)" AT %I2314.6 : Bool;   // SPARE SAFETY INPUT
   "Carrier_39_SpareSafetyInput(2_7)" AT %I2314.7 : Bool;   // SPARE SAFETY INPUT
   "Carrier_39_Slot3_SafetyOutput" AT %IW2315 : Word;   // SLOT 3 SAFETY OUTPUT WORD
   "Carrier_39_Crash_Detect_OK" AT %I2315.0 : Bool;   // CARRIER CRASH DETECT
   "Carrier_39_SpareSafetyOutput(3_1)" AT %I2315.1 : Bool;   // SPARE SAFETY OUTPUT
   "Carrier_39_SpareSafetyOutput(3_2)" AT %I2315.2 : Bool;   // SPARE SAFETY OUTPUT
   "Carrier_39_SpareSafetyOutput(3_3)" AT %I2315.3 : Bool;   // SPARE SAFETY OUTPUT
   "Carrier_39_SpareSafetyOutput(3_4)" AT %I2315.4 : Bool;   // SPARE SAFETY OUTPUT
   "Carrier_39_SpareSafetyOutput(3_5)" AT %I2315.5 : Bool;   // SPARE SAFETY OUTPUT
   "Carrier_39_SpareSafetyOutput(3_6)" AT %I2315.6 : Bool;   // SPARE SAFETY OUTPUT
   "Carrier_39_SpareSafetyOutput(3_7)" AT %I2315.7 : Bool;   // SPARE SAFETY OUTPUT
   "Carrier_39_Slot4_Input" AT %IW2316 : Word;   // SLOT 4 INPUT WORD
   "Carrier_39_480VPowerOn_MDCB1" AT %I2316.0 : Bool;   // 480 VAC POWER ON MDCB 1
   "Carrier_39_SpareInput(4_1)" AT %I2316.1 : Bool;   // SPARE INPUT
   "Carrier_39_SpareInput(4_2)" AT %I2316.2 : Bool;   // SPARE INPUT
   "Carrier_39_SitopSelectStatus" AT %I2316.3 : Bool;   // SITOP SELECT STATUS
   "Carrier_39_DCsupplyOnPSCB2" AT %I2316.4 : Bool;   // DC SUPPLY ON PSCB 2
   "Carrier_39_SpareInput(4_5)" AT %I2316.5 : Bool;   // SPARE INPUT
   "Carrier_39_SpareInput(4_6)" AT %I2316.6 : Bool;   // SPARE INPUT
   "Carrier_39_SpareInput(4_7)" AT %I2316.7 : Bool;   // SPARE INPUT
   "Carrier_39_PB1_ProdHoldLH" AT %I2317.0 : Bool;   // PB 1 PRODUCTION HOLD LH
   "Carrier_39_PB2_ResetLH" AT %I2317.1 : Bool;   // PB 2 RESET LH
   "Carrier_39_PB3_ProdHoldRH" AT %I2317.2 : Bool;   // PB 3 PRODUCTION HOLD RH
   "Carrier_39_PB4_ResetRH" AT %I2317.3 : Bool;   // PB 4 RESET RH
   "Carrier_39_SpareInput(4_14)" AT %I2317.4 : Bool;   // SPARE INPUT
   "Carrier_39_SpareInput(4_15)" AT %I2317.5 : Bool;   // SPARE INPUT
   "Carrier_39_SpareInput(4_16)" AT %I2317.6 : Bool;   // SPARE INPUT
   "Carrier_39_SpareInput(4_17)" AT %I2317.7 : Bool;   // SPARE INPUT
   "Carrier_39_Slot5_Output" AT %IW2318 : Word;   // SLOT 5 OUTPUT WORD
   "Carrier_39_IRD400_HMI_24VDC_ENABLE" AT %I2318.0 : Bool;   // IRD 400 PANEL HMI 24V DC POWER
   "Carrier_39_FaultLight_LH" AT %I2318.1 : Bool;   // FAULT LIGHT LH
   "Carrier_39_RunLight_LH" AT %I2318.2 : Bool;   // RUN LIGHT LH
   "Carrier_39_FaultLight_RH" AT %I2318.3 : Bool;   // FAULT LIGHT RH
   "Carrier_39_RunLight_RH" AT %I2318.4 : Bool;   // RUN LIGHT RH
   "Carrier_39_SpareOutput(5_5)" AT %I2318.5 : Bool;   // SPARE OUTPUT
   "Carrier_39_SpareOutput(5_6)" AT %I2318.6 : Bool;   // SPARE OUTPUT
   "Carrier_39_SpareOutput(5_7)" AT %I2318.7 : Bool;   // SPARE OUTPUT
   "Carrier_39_ActualSpeed" AT %IW2320 : Word;   // ACTUAL SPEED
   "Carrier_39_CarrierDriveAlarm" AT %IW2322 : Word;   // CARRIER DRIVE ALARM
   "Carrier_39_CarrierDriveWarning" AT %IW2324 : Word;   // CARRIER DRIVE WARNING
   "Carrier_40_Status" AT %IW2350 : Word;   // CARRIER STATUS WORD
   "Carrier_40_Status.0" AT %I2350.0 : Bool;   // HEARTBEAT
   "Carrier_40_Status.1" AT %I2350.1 : Bool;   // MANUAL
   "Carrier_40_Status.2" AT %I2350.2 : Bool;   // IN_AUTO
   "Carrier_40_Status.3" AT %I2350.3 : Bool;   // POSITIONING_COMPLETE
   "Carrier_40_Status.4" AT %I2350.4 : Bool;   // PRODUCTION HOLD
   "Carrier_40_Status.5" AT %I2350.5 : Bool;   // CARRIER MOVING FORWARD
   "Carrier_40_Status.6" AT %I2350.6 : Bool;   // CARRIER MOVING REVERSE
   "Carrier_40_Status.7" AT %I2350.7 : Bool;   // CARRIER FAULT
   "Carrier_40_Status.8" AT %I2351.0 : Bool;   // CRASH DETECT TRIPPED
   "Carrier_40_Status.9" AT %I2351.1 : Bool;
   "Carrier_40_Status.10" AT %I2351.2 : Bool;
   "Carrier_40_Status.11" AT %I2351.3 : Bool;
   "Carrier_40_Status.12" AT %I2351.4 : Bool;
   "Carrier_40_Status.13" AT %I2351.5 : Bool;
   "Carrier_40_Status.14" AT %I2351.6 : Bool;
   "Carrier_40_Status.15" AT %I2351.7 : Bool;
   "Carrier_40_SDCFaultCode" AT %IW2352 : Word;   // SDC FAULT CODE
   "Carrier_40_CarrierPosition" AT %ID2354 : DWord;   // CARRIER POSITION
   "Carrier_40_CarrierNumber" AT %IW2358 : Word;   // CARRIER NUMBER
   "Carrier_40_G120DControlWord" AT %IW2360 : Word;   // G120D_STW1_CONTROL
   "Carrier_40_G120DControlWord.0" AT %I2360.0 : Bool;   // Bit_00_ON
   "Carrier_40_G120DControlWord.1" AT %I2360.1 : Bool;   // Bit_01_AUS2_INH
   "Carrier_40_G120DControlWord.2" AT %I2360.2 : Bool;   // Bit_02_AUS3_STOP
   "Carrier_40_G120DControlWord.3" AT %I2360.3 : Bool;   // Bit_03_EN
   "Carrier_40_G120DControlWord.4" AT %I2360.4 : Bool;   // Bit_04_EN_RAMP
   "Carrier_40_G120DControlWord.5" AT %I2360.5 : Bool;   // Bit_05_START_RAMP
   "Carrier_40_G120DControlWord.6" AT %I2360.6 : Bool;   // Bit_06_SETPOINT
   "Carrier_40_G120DControlWord.7" AT %I2360.7 : Bool;   // Bit_07_RESET
   "Carrier_40_G120DControlWord.8" AT %I2361.0 : Bool;   // Bit_08_JOG_R
   "Carrier_40_G120DControlWord.9" AT %I2361.1 : Bool;   // Bit_09_JOG_L
   "Carrier_40_G120DControlWord.10" AT %I2361.2 : Bool;   // Bit_10_CONTR_PLC
   "Carrier_40_G120DControlWord.11" AT %I2361.3 : Bool;   // Bit_11_REVERSE
   "Carrier_40_G120DControlWord.12" AT %I2361.4 : Bool;   // Bit_12_BRAKE_RELEASE
   "Carrier_40_G120DControlWord.13" AT %I2361.5 : Bool;   // Bit_13_DDS
   "Carrier_40_G120DControlWord.14" AT %I2361.6 : Bool;   // Bit_14_DO0
   "Carrier_40_G120DControlWord.15" AT %I2361.7 : Bool;   // Bit_15_DO1
   "Carrier_40_G120DStatusWord" AT %IW2362 : Word;   // G120D_ZSW1_STATUS
   "Carrier_40_G120DStatusWord.0" AT %I2362.0 : Bool;   // Bit_00_READY_RUN
   "Carrier_40_G120DStatusWord.1" AT %I2362.1 : Bool;   // Bit_01_READY_ON
   "Carrier_40_G120DStatusWord.2" AT %I2362.2 : Bool;   // Bit_02_ENABLE
